                                       REGION "BUTTON SELECTED"
                                           #animate := "Animate Bool"(colorTrue := "BgLTe",
                                                                      colorFalse := #animate,
                                                                      evalSignal := #settings.kp8.btnSelState[#i]);
                                       END_REGION

                                       REGION "BUTTON UP/DOWN"
                                           #animate := "Animate Bool"(colorTrue := "BgDTe",
                                                                      colorFalse := #animate,
                                                                      evalSignal := #btnPress);
                                       END_REGION
                                   END_IF;
                               END_REGION

                               REGION "SAVE ANIMATION"
                                   #settings.kp8.buttons[#i].animate := #animate;
                               END_REGION

                           END_REGION

                       END_IF;
                   END_REGION

               END_FOR;
           END_REGION

       END_REGION

   END_REGION

   REGION "DRAW KP8 BUTTON LABELS"
       IF #reset THEN
           #settings.kp8.buttons[1].label := wstring#'6';
           #settings.kp8.buttons[2].label := wstring#'4';
           #settings.kp8.buttons[3].label := wstring#'2';
           #settings.kp8.buttons[5].label := wstring#'5';
           #settings.kp8.buttons[6].label := wstring#'3';
           #settings.kp8.buttons[7].label := wstring#'1';
       END_IF;
   END_REGION

   REGION "CHANGE DETECTION"
       #oldSelState := #settings.kp8.btnSelState;
   END_REGION
END_FUNCTION_BLOCK

FUNCTION_BLOCK "Buffer Log: Part Requests"   // FB22, SCL
{ S7_Optimized_Access := 'TRUE' }
VERSION : 0.1
   VAR_INPUT
      stations : "Stations";
   END_VAR
   VAR_IN_OUT
      logBuffer : "Part Req Log";
      logFlag : Int;
   END_VAR
   VAR
      clpsLogTime : Real;
      old : Struct
         ordered : "Station Old Presses";
         requested : "Station Old Presses";
      END_STRUCT;
      pLogBuffer : Int;
      rt : "Runtime Data";
   END_VAR
   VAR_TEMP
      address : Int;
      btnCount : Int;
      clpsFlag : Bool;
      i : Int;
      j : Int;
      oldPartOrdered : Bool;
      oldPartReq : Bool;
      partOrdered : Bool;
      partReq : Bool;
      stnCount : Int;
      readTimeRetVal : Int;
      blankRow : "Part Req Log Row";
   END_VAR
   VAR CONSTANT
      clpsItrvl : Real := 2.0;
      fulfilled : Int := 3;
      ordered : Int := 2;
      requested : Int := 1;
   END_VAR
BEGIN
   REGION "RUNTIME CALL"
       #rt.elapsed := RUNTIME(#rt.mem);
       #rt.asReal := LREAL_TO_REAL(#rt.elapsed);
   END_REGION

   REGION "COPY TO LOCAL"
       #btnCount := "ptsPerStn";
       #stnCount := "stnCount";
   END_REGION

   REGION "FOR EACH STATION"
       FOR #i := 0 TO #stnCount DO

           REGION "FOR EACH BUTTON"
               FOR #j := 0 TO #btnCount DO

                   REGION "COPY TO LOCAL"
                       #partOrdered := #stations.me[#i].partOrdered[#j];
                       #partReq := #stations.me[#i].partRequested[#j];
                       #oldPartOrdered := #old.ordered.me[#i,#j];
                       #oldPartReq := #old.requested.me[#i,#j];
                   END_REGION;

                   REGION "CALCULATE ADDRESS"
                       #address := (#i + 1) * 10 + #j + 1;
                   END_REGION

                   REGION "ON PART REQUEST RISING EDGE"
                       IF #partReq AND NOT #oldPartReq THEN

                           REGION "LOG ENTRY"
                               #logBuffer.me[#pLogBuffer] := "Buffer Part Req Log Row: Generate"(address := #address,
                                                                                        type := #requested);
                           END_REGION

                           REGION "INCREMENT POINTER"
                               #pLogBuffer += 1;
                           END_REGION

                       END_IF;
                   END_REGION

                   REGION "ON PART ORDERED RISING EDGE"
                       IF #partOrdered AND NOT #oldPartOrdered THEN

                           REGION "REQUEST TYPE"
                               #logBuffer.me[#pLogBuffer] := "Buffer Part Req Log Row: Generate"(address := #address,
                                                                                                 type := #ordered);
                           END_REGION

                           REGION "INCREMENT POINTER"
                               #pLogBuffer += 1;
                           END_REGION

                       END_IF;
                   END_REGION

                   REGION "ON PART REQUEST FALLING EDGE"
                       IF NOT #partReq AND #oldPartReq THEN

                           REGION "REQUEST TYPE"
                               #logBuffer.me[#pLogBuffer] := "Buffer Part Req Log Row: Generate"(
                                   address := #address,
                                   type := #fulfilled
                               );
                           END_REGION

                           REGION "INCREMENT POINTER"
                               #pLogBuffer += 1;
                           END_REGION

                       END_IF;
                   END_REGION

                   REGION "SAVE FOR CHANGE DETECTION"
                       #old.requested.me[#i, #j] := #partReq;
                       #old.ordered.me[#i, #j] := #partOrdered;
                   END_REGION

               END_FOR;
           END_REGION

       END_FOR;
   END_REGION

   REGION "SEND TO HMI"

       REGION "ON ENTRY IN BUFFER"
           IF #logBuffer.me[0].address <> 0 THEN

               REGION "TIMER"
                   #clpsLogTime += #rt.asReal;
                   IF #clpsLogTime >= #clpsItrvl THEN
                       #clpsLogTime := 0.0;
                       #clpsFlag := TRUE;
                   END_IF;
               END_REGION

               REGION "EXECUTE COLLAPSE"
                   IF #clpsFlag THEN

                       REGION "MOVE BUFFER UP ONE POSITION"
                           FOR #i := 0 TO 98 DO
                               #logBuffer.me[#i] := #logBuffer.me[#i + 1];
                           END_FOR;
                       END_REGION

                       REGION "DELETE LAST ROW"
                           #logBuffer.me[99] := #blankRow;
                       END_REGION

                       REGION "FLAG FOR HMI"
                           #logFlag += 1;
                           IF #logFlag > 9 THEN
                               #logFlag := 0;
                           END_IF;
                       END_REGION

                       REGION "DECREMENT POINTER"
                           #pLogBuffer -= 1;
                       END_REGION

                   END_IF;
               END_REGION

           END_IF;
       END_REGION

   END_REGION

   REGION "RESET TIMER"
       IF #logBuffer.me[0].address = 0 THEN
           #clpsLogTime := 0.0;
       END_IF;
   END_REGION
END_FUNCTION_BLOCK

FUNCTION_BLOCK "Enable Assignment Pair"   // FB23, SCL
{ S7_Optimized_Access := 'TRUE' }
VERSION : 0.1
   VAR_INPUT
      disable : Bool;
      enable : Bool;
   END_VAR
   VAR_IN_OUT
      value : WString;
      assignAnimate : USInt;
      ioFieldAnimate : USInt;
   END_VAR
   VAR
      old : Struct
         disabled : Bool;
         enabled : Bool;
      END_STRUCT;
   END_VAR
BEGIN
   REGION "DISABLED"    
       IF #disable THEN
           #value := wstring#'';
           #assignAnimate := "disabled";
           #ioFieldAnimate := "disabled";
       END_IF;
   END_REGION

   REGION "ENABLED"
           IF #enable THEN
               #assignAnimate := "BgGray";
               #ioFieldAnimate := "BgWh";
           END_IF;
   END_REGION
END_FUNCTION_BLOCK

FUNCTION_BLOCK "Assign Button Parameters"   // FB24, SCL
{ S7_Optimized_Access := 'TRUE' }
VERSION : 0.1
   VAR_INPUT
      settings : "Settings";
   END_VAR
   VAR_IN_OUT
      stations : "Stations";
   END_VAR
   VAR
      old : Struct
         allotted : Bool;
         critical : Bool;
         pn : Bool;
      END_STRUCT;
   END_VAR
   VAR_TEMP
      assign : Bool;
      btn : Struct
         allotted : Bool;
         critical : Bool;
         pn : Bool;
      END_STRUCT;
      btnSelected : Bool;
      i : Int;
      j : Int;
      partNumber : WString;
      stnSelected : Bool;
      timerReal : Real;
   END_VAR
BEGIN
   REGION "COPY TO LOCACL"
       #btn.allotted := #settings.alotted.assign.actuate;
       #btn.critical := #settings.critical.assign.actuate;
       #btn.pn := #settings.partNumber.assign.actuate;
   END_REGION

   REGION "ASSIGNMENT PULSE"
       #assign := (#btn.allotted AND NOT #old.allotted)
                   OR (#btn.critical AND NOT #old.critical)
                   OR (#btn.pn AND NOT #old.pn);
   END_REGION

   REGION "ON ASSIGNMENT PULSE"
       IF #assign THEN
           REGION "PROCESS VARIABLE"

               REGION "PART NUMBER"
                   IF #btn.pn THEN
                       #partNumber := #settings.partNumber.ioField.value;
                   END_IF;
               END_REGION

               REGION "CRITICAL TIME"
                   IF #btn.critical THEN
                       #timerReal := "WString Timer to Real"(#settings.critical.ioField.value);
                   END_IF;
               END_REGION

               REGION "ALLOTTED TIME"
                   IF #btn.allotted THEN
                       #timerReal := "WString Timer to Real"(#settings.alotted.ioField.value);
                   END_IF;
               END_REGION

           END_REGION

           REGION "FOR EACH STATION"
               FOR #i := 0 TO "stnCount" DO

                   REGION "COPY TO LOCAL"
                       #stnSelected := #stations.me[#i].settings.selected;
                   END_REGION

                   REGION "ON SELECTED STATION"
                       IF #stnSelected THEN

                           REGION "FOR EACH BUTTON"
                               FOR #j := 0 TO "ptsPerStn" DO

                                   REGION "COPY TO LOCAL"
                                       #btnSelected := #stations.me[#i].settings.btnSelection[#j];
                                   END_REGION

                                   REGION "ON SELECTED BUTTON"
                                       IF #btnSelected THEN

                                           REGION "ASSIGN PART NUMBER"
                                               IF #btn.pn THEN
                                                   #stations.me[#i].partNumbers[#j] := #partNumber;
                                               END_IF;
                                           END_REGION

                                           REGION "ASSIGN ALLOTTED TIME"
                                               IF #btn.allotted THEN
                                                   #stations.me[#i].presetTime.allotted[#j] := #timerReal;
                                               END_IF;
                                           END_REGION

                                           REGION "ASSIGN CRITICAL TIME"
                                               IF #btn.critical THEN
                                                   #stations.me[#i].presetTime.critical[#j] := #timerReal;
                                               END_IF;
                                           END_REGION

                                       END_IF;
                                   END_REGION

                               END_FOR;
                           END_REGION

                       END_IF;
                   END_REGION

               END_FOR;
           END_REGION

       END_IF;
   END_REGION

   REGION "CHANGE DETECTION"
       #old := #btn;
   END_REGION
END_FUNCTION_BLOCK

FUNCTION_BLOCK "Animate: PN & Timers"   // FB25, SCL
{ S7_Optimized_Access := 'TRUE' }
VERSION : 0.1
   VAR_INPUT
      stations : "Stations";
   END_VAR
   VAR_IN_OUT
      settings : "Settings";
   END_VAR
   VAR
      instPNEntEnable : "Enable Assignment Pair";
      instAlltEntEnable : "Enable Assignment Pair";
      instCrtEntEnable : "Enable Assignment Pair";
   END_VAR
   VAR_TEMP
      animate : USInt;
      disable : Bool;
      enable : Bool;
      selBtnCount : Int;
      selStnCount : Int;
   END_VAR
BEGIN
   REGION "COPY TO LOCAL"
       #selBtnCount := #settings.kp8.selCount;
       #selStnCount := #settings.stations.selCount;
   END_REGION

   REGION "ENABLE/DISABLE FOR PN AND TIMERS"

       REGION "SET DISABLE"
           IF #selStnCount = 0 OR #selBtnCount = 0 THEN
               #disable := TRUE;
               #enable := FALSE;
           END_IF;
       END_REGION

       REGION "SET ENABLE"
           IF #selStnCount <> 0 AND #selBtnCount <> 0 THEN
               #disable := FALSE;
               #enable := TRUE;
           END_IF;
       END_REGION

   END_REGION

   REGION "PN ANIMATION FUNCTIONS"
       #animate := #settings.partNumber.assign.animate;
       #instPNEntEnable(disable := #disable,
                        enable := #enable,
                        value := #settings.partNumber.ioField.value,
                        assignAnimate := #animate,
                        ioFieldAnimate := #settings.partNumber.ioField.animate);
       #animate := "Animate Bool"(colorTrue := "BgLGr",
                                  colorFalse := #animate,
                                  evalSignal := #settings.partNumber.assign.actuate);
       #settings.partNumber.assign.animate := #animate;
   END_REGION

   REGION "ALLOTTED TIME ANIMATION FUNCTIONS"
       #animate := #settings.alotted.assign.animate;
       #instAlltEntEnable(disable := #disable,
                          enable := #enable,
                          value := #settings.alotted.ioField.value,
                          assignAnimate := #animate,
                          ioFieldAnimate := #settings.alotted.ioField.animate);
       #animate := "Animate Bool"(colorTrue := "BgLGr",
                                  colorFalse := #animate,
                                  evalSignal := #settings.alotted.assign.actuate);
       #settings.alotted.assign.animate := #animate;
   END_REGION

   REGION "CRITICAL TIME ANIMATION FUNCTIONS"
       #animate := #settings.critical.assign.animate;
       #instCrtEntEnable(disable := #disable,
                         enable := #enable,
                         value := #settings.critical.ioField.value,
                         assignAnimate := #animate,
                         ioFieldAnimate := #settings.critical.ioField.animate);
       #animate := "Animate Bool"(colorTrue := "BgLGr",
                                  colorFalse := #animate,
                                  evalSignal := #settings.critical.assign.actuate);
       #settings.critical.assign.animate := #animate;
   END_REGION
END_FUNCTION_BLOCK

FUNCTION_BLOCK "Global to Sim"   // FB26, SCL
{ S7_Optimized_Access := 'TRUE' }
VERSION : 0.1
   VAR_INPUT
      stations : "Stations";
   END_VAR
   VAR_IN_OUT
      simStations : "Simulated Stations";
   END_VAR
   VAR
      old : Struct
         nextGrp : Bool;
         prevGrp : Bool;
      END_STRUCT;
   END_VAR
   VAR_TEMP
      animate : USInt;
      btnCount : Int;
      currentBtn : Bool;
      dzLabel : WString;
      firstStn : Int;
      i : Int;
      intBox : Int;
      j : Int;
      kp8Color : DWord;
      label : WString;
      oldBtn : Bool;
      pSim : Int;
      pStn : Int;
      simKP8Count : Int;
      stnCount : Int;
   END_VAR
   VAR CONSTANT
      space : WString := WSTRING#' ';
      lead0 : WString := WSTRING#'0';
      volvo16 : WString := WSTRING#'VOLVO 16';
   END_VAR
BEGIN
   REGION "COPY TO LOCAL"
       #btnCount := "ptsPerStn";
       #firstStn := #simStations.firstStn;
       #stnCount := "stnCount";
       #simKP8Count := "simKP8Count";
   END_REGION

   REGION "RESOLVE STATION POINTER"

       REGION "PROCESS NEXT GROUP PRESS"

           REGION "COPY TO LOCAL"
               #currentBtn := #simStations.down.actuate;
               #oldBtn := #old.nextGrp;
           END_REGION

           REGION "FALLING EDGE OF NEXT GROUP"
               IF NOT #currentBtn AND #oldBtn THEN

                   REGION "INCREMENT FIRST STATION"
                       #firstStn += #simKP8Count;
                   END_REGION

                   REGION "UPPER LIMIT ROLL OVER"
                       IF #firstStn > #stnCount THEN
                           #firstStn -= #stnCount + 1;
                       END_IF;
                   END_REGION

               END_IF;
           END_REGION

           REGION "NEXT GROUP CHANGE DETECTION"
               #old.nextGrp := #currentBtn;
           END_REGION

       END_REGION

       REGION "PROCESS PREVIOUS GROUP PRESS"

           REGION "COPY TO LOCAL"
               #currentBtn := #simStations.up.actuate;
               #oldBtn := #old.prevGrp;
           END_REGION

           REGION "FALLING EDGE OF PREVIOUS GROUP"
               IF NOT #currentBtn AND #oldBtn THEN

                   REGION "DECREMENT FIRST STATION"
                       #firstStn -= #simKP8Count;
                   END_REGION

                   REGION "LOWER LIMIT ROLL OVER"
                       IF #firstStn < 0 THEN
                           #firstStn += #stnCount + 1;
                       END_IF;
                   END_REGION

               END_IF;
           END_REGION

           REGION "PREVIOUS GROUP CHANGE DETECTION"
               #old.prevGrp := #currentBtn;
           END_REGION

       END_REGION

   END_REGION

   REGION "FOR EACH BUTTON"
       FOR #i := 0 TO 11 DO

           REGION "CALCULATE POINTER"
               #pStn := #i + #firstStn;
               #pSim := #i;
           END_REGION

           REGION "UPPER LIMIT ROLL OVER"
               IF #pStn > #stnCount THEN
                   #pStn := #firstStn + #i - #stnCount - 1;
               END_IF;
           END_REGION

           REGION "COPY TO LOCAL"
               #kp8Color := #stations.me[#pStn].kp8Out;
           END_REGION

           REGION "LABEL STATIONS"

               REGION "DETERMINE LINE LABEL"
                   #label := #stations.me[#pStn].line;
                   IF #label = #volvo16 THEN
                       #label := WSTRING#'V16';
                   END_IF;
               END_REGION

               REGION "DETERMINE DROP ZONE LABEL"
                   #intBox := USINT_TO_INT(#stations.me[#pStn].dropZone);
                   IF #intBox <= 9 THEN
                       #dzLabel := CONCAT_WSTRING(IN1 := #lead0,
                                                  IN2 := "Strip Sign"(INT_TO_WSTRING(#intBox)));
                   END_IF;
                   IF #intBox >= 10 THEN
                       #dzLabel := "Strip Sign"(INT_TO_WSTRING(#intBox));
                   END_IF;
               END_REGION

               REGION "WRITE LABEL"
                   #label := CONCAT_WSTRING(IN1 := #label,
                                            IN2 := #space,
                                            IN3 := #dzLabel);
                   #simStations.me[#pSim].stn.label := #label;
               END_REGION

           END_REGION

           REGION "ANIMATE STATION LABEL"
               #simStations.me[#pSim].stn.animate := "BgGray";
           END_REGION

           REGION "FOR EACH BUTTON"
               FOR #j := 0 TO #btnCount DO

                   REGION "COLOR BUTTONS"
                       #animate := "KP8 Color to Sim Animation"(kp8Color := #kp8Color,
                                                                btnNumber := #j);
                       #simStations.me[#pSim].btn.animate[#j] := #animate;
                   END_REGION

                   REGION "WRITE BUTTON LABELS"
                       #intBox := "Pointer Calc: KP8 Labels"(#j);
                       #label := "Strip Sign"(INT_TO_WSTRING(#intBox));
                       #simStations.me[#pSim].btn.labels[#j] := #label;
                   END_REGION

               END_FOR;
           END_REGION

       END_FOR;
   END_REGION

   REGION "SAVE FIRST STATION"
       #simStations.firstStn := #firstStn;
   END_REGION

   REGION "ANIMATE NEXT GROUP PRESS"
       #simStations.down.animate := "Animate Bool"(colorTrue := "BgLGr",
                                                   colorFalse := "BgGray",
                                                   evalSignal := #simStations.down.actuate);
   END_REGION

   REGION "ANIMATE PREV GROUP PARESS"
       #simStations.up.animate := "Animate Bool"(colorTrue := "BgLGr",
                                                 colorFalse := "BgGray",
                                                 evalSignal := #simStations.up.actuate);
   END_REGION
END_FUNCTION_BLOCK

FUNCTION_BLOCK "HMI: Network Health"   // FB31, SCL
{ S7_Optimized_Access := 'TRUE' }
VERSION : 0.1
   VAR_IN_OUT
      ioSystemData : Array[1.."USERDIAG_IO_SYSTEMS_UPPER_LIM"] of "UserDiag_typeIOSystem";
      netHealthScreen : "Network Health Screen";
   END_VAR
   VAR_TEMP
      i : Int;
      animate : Struct
         ok : USInt;
         faulty : USInt;
         lostConn : USInt;
         disabled : USInt;
         problem : USInt;
         wasFaulty : USInt;
         wasLost : USInt;
         wasDisabled : USInt;
         problemGone : USInt;
      END_STRUCT;
   END_VAR
   VAR CONSTANT
      statOk : USInt := 1;
   END_VAR
BEGIN
   #animate.ok := "BgDGr";

   FOR #i := 1 TO "pnioDeviceCount" DO
       #netHealthScreen.pnioDevices[#i].label := #ioSystemData[1].devices[#i].name;
       CASE #ioSystemData[1].devices[#i].state OF
           #statOk:
               #netHealthScreen.pnioDevices[#i].animate := #animate.ok;
           ELSE 
               ;
       END_CASE;
   END_FOR;
END_FUNCTION_BLOCK

FUNCTION_BLOCK "Table Navigatio"   // FB34, SCL
{ S7_Optimized_Access := 'TRUE' }
VERSION : 0.1
   VAR_INPUT
      maxRows : DInt;
      visRows : DInt;
      offset : DInt;
      trigger : Bool;
   END_VAR
   VAR_IN_OUT
      r1 : DInt;
      rowIndices : Array[0..#maxOutRows] of DInt;
   END_VAR
   VAR
      old : Struct
         trigger : Bool := false;
      END_STRUCT;
   END_VAR
   VAR_TEMP
      i : DInt;
      output : Array[0..#maxOutRows] of DInt;
      thisIndex : DInt;
      newR1 : DInt;
   END_VAR
   VAR CONSTANT
      maxOutRows : DInt := 99;
   END_VAR
BEGIN
   IF #trigger AND NOT #old.trigger THEN

       FOR #i := 0 TO #maxOutRows DO
           #output[#i] := -1;
       END_FOR;

       IF #offset > -1000 THEN

           #newR1 := #r1 + #offset;

           IF #newR1 < 0 THEN
               #newR1 := #newR1 + #maxRows;
           END_IF;

           IF #newR1 > #maxRows THEN
               #newR1 := #newR1 - #maxRows;
           END_IF;

       END_IF;

       IF #offset = -1000 THEN
           #newR1 := 0;
       END_IF;

       IF #offset = - 2000 THEN
           #newR1 := #maxRows - #visRows;
       END_IF;

       FOR #i := 0 TO #visRows - 1 DO
           #thisIndex := #newR1 + #i;
           IF #thisIndex < 0 THEN
               #thisIndex := #thisIndex + #maxRows;
           END_IF;
           IF #thisIndex >= #maxRows THEN
               #thisIndex := #thisIndex - #maxRows;
           END_IF;
           #output[#i] := #thisIndex;
       END_FOR;

       #rowIndices := #output;
       #r1 := #newR1;

   END_IF;

   #old.trigger := #trigger;
END_FUNCTION_BLOCK

FUNCTION_BLOCK "KP8 Driver"   // FB101, SCL
{ S7_Optimized_Access := 'FALSE' }
VERSION : 0.1
   VAR_INPUT
      btnIn : Byte;   // byte that contains input data from kp8 buttons
      hardInit : Bool;   // initializes function. can be used for reset
      softInit : Bool;
      btn0Activate : Bool;   // true for on, false for off
      btn0Mode : Bool;   // true for maintained, false for momentary
      btn0Group : Int;
      btn0Flash : Bool;
      btn0ColorOn1 : String[10];   // enter: red OR green OR blue OR yellow OR white OR off
      btn0ColorOn2 : String[10];
      btn0ColorOff : String[10];   // enter: red OR green OR blue OR yellow OR white OR off
      btn1Activate : Bool;   // true for on, false for off
      btn1Mode : Bool;   // true for maintained, false for momentary
      btn1Group : Int;
      btn1Flash : Bool;
      btn1ColorOn1 : String[10];   // enter: red OR green OR blue OR yellow OR white OR off
      btn1ColorOn2 : String[10];
      btn1ColorOff : String[10];   // enter: red OR green OR blue OR yellow OR white OR off
      btn2Activate : Bool;   // true for on, false for off
      btn2Mode : Bool;   // true for maintained, false for momentary
      btn2Group : Int;
      btn2Flash : Bool;
      btn2ColorOn1 : String[10] := '';   // enter: red OR green OR blue OR yellow OR white OR off
      btn2ColorOn2 : String[10];
      btn2ColorOff : String[10];   // enter: red OR green OR blue OR yellow OR white OR off
      btn3Activate : Bool;   // true for on, false for off
      btn3Mode : Bool;   // true for maintained, false for momentary
      btn3Group : Int;
      btn3Flash : Bool;
      btn3ColorOn1 : String[10];   // enter: red OR green OR blue OR yellow OR white OR off
      btn3ColorOn2 : String[10];
      btn3ColorOff : String[10];   // enter: red OR green OR blue OR yellow OR white OR off
      btn4Activate : Bool;   // true for on, false for off
      btn4Mode : Bool;   // true for maintained, false for momentary
      btn4Group : Int;
      btn4Flash : Bool;
      btn4ColorOn1 : String[10];   // enter: red OR green OR blue OR yellow OR white OR off
      btn4ColorOn2 : String[10];
      btn4ColorOff : String[10];   // enter: red OR green OR blue OR yellow OR white OR off
      btn5Activate : Bool;   // true for on, false for off
      btn5Mode : Bool;   // true for maintained, false for momentary
      btn5Group : Int;
      btn5Flash : Bool;
      btn5ColorOn1 : String[10];   // enter: red OR green OR blue OR yellow OR white OR off
      btn5ColorOn2 : String[10];
      btn5ColorOff : String[10];   // enter: red OR green OR blue OR yellow OR white OR off
      btn6Activate : Bool;   // true for on, false for off
      btn6Mode : Bool;   // true for maintained, false for momentary
      btn6Group : Int;
      btn6Flash : Bool;
      btn6ColorOn1 : String[10];   // enter: red OR green OR blue OR yellow OR white OR off
      btn6ColorOn2 : String[10];
      btn6ColorOff : String[10];   // enter: red OR green OR blue OR yellow OR white OR off
      btn7Activate : Bool;   // true for on, false for off
      btn7Mode : Bool;   // true for maintained, false for momentary
      btn7Group : Int;
      btn7Flash : Bool;
      btn7ColorOn1 : String[10];   // enter: red OR green OR blue OR yellow OR white OR off
      btn7ColorOn2 : String[10];
      btn7ColorOff : String[10];   // enter: red OR green OR blue OR yellow OR white OR off
   END_VAR
   VAR_OUTPUT
      btnStatesOut : Array[0..7] of Bool;   // the output array represents the state of button presses
      btnColorsOut : DWord;
   END_VAR
   VAR
      mask : Byte;
      btnInInt : Byte;
      btnEval : Byte;
      i1 : Int;
      i2 : Int;
      btnActivateInt : Array[0..7] of Bool;
      btnClrMskOffInt : Array[0..7] of DWord;
      btnClrMskOn1Int : Array[0..7] of DWord;
      btnClrMskOn2Int : Array[0..7] of DWord;
      btnClrOffInt : Array[0..7] of String[10];
      btnClrOn1Int : Array[0..7] of String[10];
      btnClrOn2Int : Array[0..7] of String[10];
      btnColors : DWord;
      btnInArrayNew : Array[0..7] of Bool;
      btnInArrayOld : Array[0..7] of Bool;
      btnStateArrayInt : Array[0..7] of Bool;
      btnModeInt : Array[0..7] of Bool;
      btnFlashInt : Array[0..7] of Bool;
      btnGroup : Array[0..7] of Int;
   END_VAR
   VAR CONSTANT
      btnMskRed : DWord := dw#16#0100_0000;
      btnMskGreen : DWord := dw#16#0001_0000;
      btnMskBlue : DWord := dw#16#000_0100;
      btnMskYellow : DWord := dw#16#0101_0000;
      btnMskWhite : DWord := dw#16#0101_0100;
      btnMskBlack : DWord := dw#16#FEFE_FEFF;
      initBtnColors : DWord := dw#16#0000_0000;
   END_VAR
BEGIN
   REGION "ALL INITS"
       IF #hardInit OR #softInit THEN

           REGION "CLEAR OUTPUT COLORS"
               #btnColors := #initBtnColors;
           END_REGION

           REGION "TRANSFER PARAMETERS TO INTERNAL ARRAYS"

               REGION "BUTTON 0"
                   #btnActivateInt[0] := #btn0Activate;
                   #btnModeInt[0] := #btn0Mode;
                   #btnGroup[0] := #btn0Group;
                   #btnClrOn1Int[0] := #btn0ColorOn1;
                   #btnClrOn2Int[0] := #btn0ColorOn2;
                   #btnClrOffInt[0] := #btn0ColorOff;
               END_REGION

               REGION "BUTTON 1"
                   #btnActivateInt[1] := #btn1Activate;
                   #btnModeInt[1] := #btn1Mode;
                   #btnGroup[1] := #btn1Group;
                   #btnClrOn1Int[1] := #btn1ColorOn1;
                   #btnClrOn2Int[1] := #btn1ColorOn2;
                   #btnClrOffInt[1] := #btn1ColorOff;
               END_REGION

               REGION "BUTTON 2"
                   #btnActivateInt[2] := #btn2Activate;
                   #btnModeInt[2] := #btn2Mode;
                   #btnGroup[2] := #btn2Group;
                   #btnClrOn1Int[2] := #btn2ColorOn1;
                   #btnClrOn2Int[2] := #btn2ColorOn2;
                   #btnClrOffInt[2] := #btn2ColorOff;
               END_REGION

               REGION "BUTTON 3"
                   #btnActivateInt[3] := #btn3Activate;
                   #btnModeInt[3] := #btn3Mode;
                   #btnGroup[3] := #btn3Group;
                   #btnClrOn1Int[3] := #btn3ColorOn1;
                   #btnClrOn2Int[3] := #btn3ColorOn2;
                   #btnClrOffInt[3] := #btn3ColorOff;
               END_REGION

               REGION "BUTTON 4"
                   #btnActivateInt[4] := #btn4Activate;
                   #btnModeInt[4] := #btn4Mode;
                   #btnGroup[4] := #btn4Group;
                   #btnClrOn1Int[4] := #btn4ColorOn1;
                   #btnClrOn2Int[4] := #btn4ColorOn2;
                   #btnClrOffInt[4] := #btn4ColorOff;
               END_REGION

               REGION "BUTTON 5"
                   #btnActivateInt[5] := #btn5Activate;
                   #btnModeInt[5] := #btn5Mode;
                   #btnGroup[5] := #btn5Group;
                   #btnClrOn1Int[5] := #btn5ColorOn1;
                   #btnClrOn2Int[5] := #btn5ColorOn2;
                   #btnClrOffInt[5] := #btn5ColorOff;
               END_REGION

               REGION "BUTTON 6"
                   #btnActivateInt[6] := #btn6Activate;
                   #btnModeInt[6] := #btn6Mode;
                   #btnGroup[6] := #btn6Group;
                   #btnClrOn1Int[6] := #btn6ColorOn1;
                   #btnClrOn2Int[6] := #btn6ColorOn2;
                   #btnClrOffInt[6] := #btn6ColorOff;
               END_REGION

               REGION "BUTTON 7"
                   #btnActivateInt[7] := #btn7Activate;
                   #btnModeInt[7] := #btn7Mode;
                   #btnGroup[7] := #btn7Group;
                   #btnClrOn1Int[7] := #btn7ColorOn1;
                   #btnClrOn2Int[7] := #btn7ColorOn2;
                   #btnClrOffInt[7] := #btn7ColorOff;
               END_REGION

           END_REGION

           REGION "RECOLOR BUTTON MASKS"
               FOR #i1 := 0 TO 7 DO

                   REGION "ON COLOR 1"
                       IF (#btnClrOn1Int[#i1] = 'red') THEN
                           #btnClrMskOn1Int[#i1] := SHL(IN := #btnMskRed, N := INT_TO_ULINT(#i1));
                       ELSIF (#btnClrOn1Int[#i1] = 'green') THEN
                           #btnClrMskOn1Int[#i1] := SHL(IN := #btnMskGreen, N := INT_TO_ULINT(#i1));
                       ELSIF (#btnClrOn1Int[#i1] = 'blue') THEN
                           #btnClrMskOn1Int[#i1] := SHL(IN := #btnMskBlue, N := INT_TO_ULINT(#i1));
                       ELSIF (#btnClrOn1Int[#i1] = 'yellow') THEN
                           #btnClrMskOn1Int[#i1] := SHL(IN := #btnMskYellow, N := INT_TO_ULINT(#i1));
                       ELSIF (#btnClrOn1Int[#i1] = 'white') THEN
                           #btnClrMskOn1Int[#i1] := SHL(IN := #btnMskWhite, N := INT_TO_ULINT(#i1));
                       ELSIF (#btnClrOn1Int[#i1] = 'off') THEN
                           #btnClrMskOn1Int[#i1] := 0;
                       END_IF;
                   END_REGION

                   REGION "ON COLOR 2"
                       IF (#btnClrOn2Int[#i1] = 'red') THEN
                           #btnClrMskOn2Int[#i1] := SHL(IN := #btnMskRed, N := INT_TO_ULINT(#i1));
                       ELSIF (#btnClrOn2Int[#i1] = 'green') THEN
                           #btnClrMskOn2Int[#i1] := SHL(IN := #btnMskGreen, N := INT_TO_ULINT(#i1));
                       ELSIF (#btnClrOn2Int[#i1] = 'blue') THEN
                           #btnClrMskOn2Int[#i1] := SHL(IN := #btnMskBlue, N := INT_TO_ULINT(#i1));
                       ELSIF (#btnClrOn2Int[#i1] = 'yellow') THEN
                           #btnClrMskOn2Int[#i1] := SHL(IN := #btnMskYellow, N := INT_TO_ULINT(#i1));
                       ELSIF (#btnClrOn2Int[#i1] = 'white') THEN
                           #btnClrMskOn2Int[#i1] := SHL(IN := #btnMskWhite, N := INT_TO_ULINT(#i1));
                       ELSIF (#btnClrOn2Int[#i1] = 'off') THEN
                           #btnClrMskOn2Int[#i1] := 0;
                       END_IF;
                   END_REGION

                   REGION "OFF COLOR"
                       IF (#btnClrOffInt[#i1] = 'red') THEN
                           #btnClrMskOffInt[#i1] := SHL(IN := #btnMskRed, N := INT_TO_ULINT(#i1));
                       ELSIF (#btnClrOffInt[#i1] = 'green') THEN
                           #btnClrMskOffInt[#i1] := SHL(IN := #btnMskGreen, N := INT_TO_ULINT(#i1));
                       ELSIF (#btnClrOffInt[#i1] = 'blue') THEN
                           #btnClrMskOffInt[#i1] := SHL(IN := #btnMskBlue, N := INT_TO_ULINT(#i1));
                       ELSIF (#btnClrOffInt[#i1] = 'yellow') THEN
                           #btnClrMskOffInt[#i1] := SHL(IN := #btnMskYellow, N := INT_TO_ULINT(#i1));
                       ELSIF (#btnClrOffInt[#i1] = 'white') THEN
                           #btnClrMskOffInt[#i1] := SHL(IN := #btnMskWhite, N := INT_TO_ULINT(#i1));
                       ELSIF (#btnClrOffInt[#i1] = 'off') THEN
                           #btnClrMskOffInt[#i1] := 0;
                       END_IF;
                   END_REGION

               END_FOR;
           END_REGION

       END_IF;
   END_REGION

   REGION "HART INIT"
       IF #hardInit THEN
           FOR #i1 := 0 TO 7 DO
               #btnStateArrayInt[#i1] := FALSE;
           END_FOR;
       END_IF;
   END_REGION


   REGION "TRANFER PARAMETERS TO ARRAYS"
       // raw pb data
       #btnInInt := #btnIn;
       // flashing modes
       #btnFlashInt[0] := #btn0Flash;
       #btnFlashInt[1] := #btn1Flash;
       #btnFlashInt[2] := #btn2Flash;
       #btnFlashInt[3] := #btn3Flash;
       #btnFlashInt[4] := #btn4Flash;
       #btnFlashInt[5] := #btn5Flash;
       #btnFlashInt[6] := #btn6Flash;
       #btnFlashInt[7] := #btn7Flash;
   END_REGION

   REGION "EVALUATE BUTTONS"
       FOR #i1 := 0 TO 7 DO

           REGION "TRANSFER BUTTON PRESSES TO ARRAY"
               #btnEval := SHR(IN := #btnInInt, N := INT_TO_ULINT(#i1));
               #btnInArrayNew[#i1] := #btnEval.%X0;
               #btnEval := b#16#0;
           END_REGION

           REGION "SET BUTTON STATE"

               REGION "BUTTON ACTIVE"
                   IF #btnActivateInt[#i1] THEN

                       REGION "MAINTAINED"
                           IF #btnModeInt[#i1] THEN

                               REGION "RISING EDGE OF PRESS"
                                   IF #btnInArrayNew[#i1] AND NOT #btnInArrayOld[#i1] THEN

                                       REGION "CHECK FOR GROUP MEMBERSHIP"
                                           FOR #i2 := 0 TO 7 DO

                                               REGION "NOT IN NULL GROUP"
                                                   IF (#btnGroup[#i2] <> 0) THEN

                                                       REGION "SKIP SELF"
                                                           IF (#i2 <> #i1) THEN

                                                               REGION "GROUPS MATCH"
                                                                   IF #btnGroup[#i1] = #btnGroup[#i2] THEN
                                                                       REGION "DEACTIVATE OTHER GROUP MEMBERS"
                                                                           #btnStateArrayInt[#i2] := FALSE;
                                                                       END_REGION

                                                                   END_IF;
                                                               END_REGION

                                                           END_IF;
                                                       END_REGION

                                                   END_IF;
                                               END_REGION

                                           END_FOR;
                                       END_REGION

                                       REGION "TOGGLE STATE"
                                           #btnStateArrayInt[#i1] := NOT #btnStateArrayInt[#i1];
                                       END_REGION

                                   END_IF;
                               END_REGION

                           END_IF;
                       END_REGION

                       REGION "MOMENTARY"
                           IF NOT #btnModeInt[#i1] THEN
                               #btnStateArrayInt[#i1] := #btnInArrayNew[#i1];
                           END_IF;
                       END_REGION

                   END_IF;
               END_REGION

               REGION "BUTTON INACTIVE"
                   IF NOT #btnActivateInt[#i1] THEN
                       #btnStateArrayInt[#i1] := FALSE;
                   END_IF;
               END_REGION

           END_REGION

           REGION "ANIMATE BUTTONS"

               REGION "BUTTON ON FLASH BIT OFF"
                   IF #btnStateArrayInt[#i1] AND NOT #btnFlashInt[#i1] THEN
                       #btnColors := #btnColors AND ROL(IN := #btnMskBlack, N := INT_TO_ULINT(#i1));
                       #btnColors := #btnColors OR #btnClrMskOn1Int[#i1];
                   END_IF;
               END_REGION

               REGION "BUTTON ON FLASH BIT ON"
                   IF #btnStateArrayInt[#i1] AND #btnFlashInt[#i1] THEN
                       #btnColors := #btnColors AND ROL(IN := #btnMskBlack, N := INT_TO_ULINT(#i1));
                       #btnColors := #btnColors OR #btnClrMskOn2Int[#i1];
                   END_IF;
               END_REGION

               REGION "BUTTON OFF"
                   IF NOT #btnStateArrayInt[#i1] THEN
                       #btnColors := #btnColors AND ROL(IN := #btnMskBlack, N := INT_TO_ULINT(#i1));
                       #btnColors := #btnColors OR #btnClrMskOffInt[#i1];
                   END_IF;
               END_REGION

           END_REGION

       END_FOR;
   END_REGION

   REGION "CHANGE DETECTION"
       #btnInArrayOld := #btnInArrayNew;
   END_REGION

   REGION "OUTPUT"
       #btnColorsOut := #btnColors;
       #btnStatesOut := #btnStateArrayInt;
   END_REGION
END_FUNCTION_BLOCK

FUNCTION "Add Leading" : WString   // FC4, SCL
{ S7_Optimized_Access := 'TRUE' }
VERSION : 0.1
   VAR_INPUT
      "Leading Character" : WChar;
      "Desired Length" : USInt;
      "String" : WString;
   END_VAR
   VAR_TEMP
      Length : Int;
      "String Box" : WString;
      Constant : WString;
   END_VAR
BEGIN
   #"String Box" := #String;
   #Length := LEN(#"String Box");

   WHILE #Length < #"Desired Length" DO
       #"String Box" := CONCAT_WSTRING(IN1 := #"Leading Character",
                                       IN2 := #"String Box");
       #Length := LEN(#"String Box");
   END_WHILE;

   #"Add Leading" := #"String Box";
END_FUNCTION

FUNCTION "Select Stations" : Void   // FC6, SCL
{ S7_Optimized_Access := 'TRUE' }
VERSION : 0.1
   VAR_INPUT
      mode : Bool;   // TRUE = select; FALSE = deselect
   END_VAR
   VAR_IN_OUT
      stations : "Stations";
   END_VAR
   VAR_TEMP
      i : Int;
      stnCount : Int;
   END_VAR
   VAR CONSTANT
      stationCount : Int := 22;
   END_VAR
BEGIN
   REGION "GET STATION COUNT"
       #stnCount := "stnCount";
   END_REGION

   REGION "SELECT STATIONS"
       FOR #i := 0 TO #stnCount DO
           #stations.me[#i].settings.selected := #mode;
       END_FOR;
   END_REGION
END_FUNCTION

FUNCTION "Dark Mode" : Void   // FC7, SCL
{ S7_Optimized_Access := 'TRUE' }
VERSION : 0.1
   VAR_IN_OUT
      animate : USInt;
   END_VAR
   VAR_TEMP
      ani : USInt;
   END_VAR
   VAR CONSTANT
      redFlashing : USInt := 12;
      invisible : USInt := 255;
      darkMode : USInt := 1;
      disabled : USInt := 254;
   END_VAR
BEGIN
   REGION "COPY TO LOCAL"
       #ani := #animate;
   END_REGION


   REGION "APPLY DARK MODE"
       CASE #ani OF
           #redFlashing, #invisible, 0, #disabled:
               #ani := #ani;
           ELSE
               #ani += #darkMode;
       END_CASE;
   END_REGION


   REGION "OUTPUT"
       #animate := #ani;
   END_REGION
END_FUNCTION

FUNCTION "Select Buttons" : Void   // FC8, SCL
{ S7_Optimized_Access := 'TRUE' }
VERSION : 0.1
   VAR_INPUT
      mode : Bool;   // TRUE = select; FALSE = deselect
   END_VAR
   VAR_IN_OUT
      stations : "Stations";
   END_VAR
   VAR_TEMP
      btnCount : Int;
      i : Int;
      j : Int;
      selected : Bool;
      stnCount : Int;
   END_VAR
   VAR CONSTANT
      buttonCount : Int := 5;
   END_VAR
BEGIN
   REGION "COPY TO LOCAL"
       #btnCount := "ptsPerStn";
       #stnCount := "stnCount";
   END_REGION

   REGION "SELECT BUTTONS"
       FOR #i := 0 TO #stnCount DO

           REGION "SELCT ALL BUTTONS ON SELECTED STATION"
               #selected := #stations.me[#i].settings.selected;
               IF #selected THEN

                   REGION "LOOP THROUGH BUTTONS"
                       FOR #j := 0 TO #btnCount DO
                           #stations.me[#i].settings.btnSelection[#j] := #mode;
                       END_FOR;
                   END_REGION

               END_IF;
           END_REGION

       END_FOR;
   END_REGION
END_FUNCTION

FUNCTION "Animate Bool" : USInt   // FC9, SCL
{ S7_Optimized_Access := 'TRUE' }
VERSION : 0.1
   VAR_INPUT
      colorTrue : USInt;
      colorFalse : USInt;
      evalSignal : Bool;
   END_VAR
   VAR_TEMP
      animate : USInt;
   END_VAR
BEGIN
   REGION "FALSE COLOR"
       IF NOT #evalSignal THEN
           #animate := #colorFalse;
       END_IF;
   END_REGION

   REGION "TRUE COLOR"
       IF #evalSignal THEN
           #animate := #colorTrue;
       END_IF;
   END_REGION

   REGION "FUNCTION RETURN"
       #"Animate Bool" := #animate;
   END_REGION
END_FUNCTION

FUNCTION "Get Part Call Row Number" : Int   // FC11, SCL
{ S7_Optimized_Access := 'TRUE' }
VERSION : 0.1
   VAR_IN_OUT
      partCall : "Part Call Screen";
   END_VAR
   VAR_TEMP
      hmiRows : Int;
      i : Int;
      selectedRow : Int;
   END_VAR
BEGIN
   REGION "GET NUMBER OF HMI ROWS"
       #hmiRows := "partReqHmiRowCount";
   END_REGION

   REGION "LOOP THROUGH HMI ROWS
       FOR #i := 0 TO #hmiRows DO

           REGION "FIND SELECTED ROW"
               IF #partCall.row[#i].pbSelection.actuate THEN
                   // selected row as int
                   #selectedRow := #i + 1;
                   EXIT;
               END_IF;
           END_REGION

       END_FOR;
   END_REGION

   REGION "RETURN ROW NUMBER"
       #"Get Part Call Row Number" := #selectedRow;
   END_REGION
END_FUNCTION

FUNCTION "Address to Station and Button" : Void   // FC12, SCL
{ S7_Optimized_Access := 'TRUE' }
VERSION : 0.1
   VAR_INPUT
      address : UInt;
   END_VAR
   VAR_OUTPUT
      station : UInt;
      button : UInt;
   END_VAR
BEGIN
   #station := #address / 10;
   #button := #address MOD 10;
END_FUNCTION

FUNCTION "Real to WString Timer" : WString   // FC14, SCL
{ S7_Optimized_Access := 'TRUE' }
VERSION : 0.1
   VAR_INPUT
      realVal : Real;
   END_VAR
   VAR CONSTANT
      msPerSec : Real := 1000.0;
   END_VAR
BEGIN
   #"Real to WString Timer" := "Time to WString"(DINT_TO_TIME(REAL_TO_DINT(#realVal * #msPerSec)));
END_FUNCTION

FUNCTION "Populate Dropzone IO Field" : WString   // FC15, SCL
{ S7_Optimized_Access := 'TRUE' }
VERSION : 0.1
   VAR_INPUT
      dzAsInt : USInt;
   END_VAR
BEGIN
   #"Populate Dropzone IO Field" := "Strip Sign"(USINT_TO_WSTRING(#dzAsInt));
END_FUNCTION

FUNCTION "Get Station Selection Number" : Void   // FC16, SCL
{ S7_Optimized_Access := 'TRUE' }
VERSION : 0.1
   VAR_INPUT
      next : Bool;   // 'next' or 'prev'
      prev : Bool;
      stations : "Stations";
   END_VAR
   VAR_IN_OUT
      selStnNumber : Int;
   END_VAR
   VAR_TEMP
      i : Int;
      stnCount : Int;
      stnSelected : Bool;
   END_VAR
BEGIN
   REGION "COPY TO LOCAL"
       #stnCount := "stnCount";
   END_REGION

   REGION "INITIALIZE INDEX"
       #i := #selStnNumber;
   END_REGION

   REGION "PREVIOUS MODE"

       REGION "DECREMENT"
           IF #prev THEN
               #i -= 1;
           END_IF;
       END_REGION

       REGION "LOW LIMIT ROLLOVER"
           IF #i < 0 THEN
               #i := #stnCount;
           END_IF;
       END_REGION

   END_REGION

   REGION "NEXT MODE"

       REGION "INCREMENT"
           IF #next THEN
               #i += 1;
           END_IF;
       END_REGION

       REGION "HIGH LIMIT ROLLOVER"
           IF #i > #stnCount THEN
               #i := 0;
           END_IF;
       END_REGION

   END_REGION

   REGION "COPY TO LOCAL"
       #stnSelected := #stations.me[#i].settings.selected;
   END_REGION

   REGION "FIND NEXT SELECTED STATION"
       WHILE NOT #stnSelected DO

           REGION "PREVIOUS MODE"

               REGION "DECREMENT"
                   IF #prev THEN
                       #i -= 1;
                   END_IF;
               END_REGION

               REGION "LOW LIMIT ROLLOVER"
                   IF #i < 0 THEN
                       #i := #stnCount;
                   END_IF;
               END_REGION

           END_REGION

           REGION "NEXT MODE"

               REGION "INCREMENT"
                   IF #next THEN
                       #i += 1;
                   END_IF;
               END_REGION

               REGION "HIGH LIMIT ROLLOVER"
                   IF #i > #stnCount THEN
                       #i := 0;
                   END_IF;
               END_REGION

           END_REGION

           REGION "SAVE WHILE CONDITION"
               #stnSelected := #stations.me[#i].settings.selected;
           END_REGION

       END_WHILE;
   END_REGION

   REGION "RETURN VALUE"
       #selStnNumber := #i;
   END_REGION
END_FUNCTION

FUNCTION "Populate Button Details" : Void   // FC17, SCL
{ S7_Optimized_Access := 'TRUE' }
VERSION : 0.1
   VAR_INPUT
      selStnNumber : Int;
      stations : "Stations";
   END_VAR
   VAR_IN_OUT
      settings : "Settings";
   END_VAR
   VAR_TEMP
      btnCount : Int;
      i : Int;
      partNumber : WString;
      pBtn : Int;
      timerWS : WString;
   END_VAR
BEGIN
   REGION "FOR EACH BUTTON"
       FOR #i := 0 TO "ptsPerStn" DO

           REGION "CALCULATE BUTTON POINTER"
               IF #i MOD 2 = 0 THEN
                   #pBtn := 7 - #i / 2;
               END_IF;
               IF #i MOD 2 <> 0 THEN
                   #pBtn := 3 - #i / 2;
               END_IF;
           END_REGION

           REGION "BUTTON LABEL"
               #settings.viewingStation.btns[#i].label.value := "Strip Sign"(INT_TO_WSTRING(#i + 1));
           END_REGION

           REGION "ALLOTTED TIME"
               #timerWS := "Real to WString Timer"(#stations.me[#selStnNumber].presetTime.allotted[#pBtn]);
               #settings.viewingStation.btns[#i].alloted.value := #timerWS;
           END_REGION

           REGION "CRITICAL TIME"
               #timerWS := "Real to WString Timer"(#stations.me[#selStnNumber].presetTime.critical[#pBtn]);
               #settings.viewingStation.btns[#i].critical.value := #timerWS;
           END_REGION

           REGION "PART NUMBER"
               #partNumber := #stations.me[#selStnNumber].partNumbers[#pBtn];
               #settings.viewingStation.btns[#i].partNumber.value := #partNumber;
           END_REGION

       END_FOR;
   END_REGION
END_FUNCTION

FUNCTION "Assign Station Parameters" : Void   // FC18, SCL
{ S7_Optimized_Access := 'TRUE' }
VERSION : 0.1
   VAR_IN_OUT
      settings : "Settings";
      stations : "Stations";
   END_VAR
   VAR_TEMP
      dzEntered : Bool;
      dzLabel : WString;
      i : Int;
      lineEntered : Bool;
      lineLabel : WString;
      stnCount : Int;
      stnSelected : Bool;
   END_VAR
BEGIN
   REGION "COPY TO LOCAL"    
       #dzEntered := #settings.viewingStation.dzData.inputFinished;
       #lineEntered := #settings.viewingStation.lineData.inputFinished;
       #stnCount := "stnCount";
   END_REGION

   REGION "ON PARAMETER ENTRY"
       IF #dzEntered OR #lineEntered THEN

           REGION "TURN OFF THE LIGHTS"
               #settings.viewingStation.dzData.inputFinished := FALSE;
               #settings.viewingStation.lineData.inputFinished := FALSE;
           END_REGION

           REGION "FOR EACH STATION"
               FOR #i := 0 TO #stnCount DO

                   REGION "COPY TO LOCAL"
                       #stnSelected := #stations.me[#i].settings.selected;
                   END_REGION

                   REGION "ON SELECTED STATION"
                       IF #stnSelected THEN

                           REGION "ON DROP ZONE INPUT"
                               IF #dzEntered THEN